(* Logix 5000 project; controller MV vendor 1 type 14 code 217 rev 31.11; software revision 31.00; part 39 of 53 *)
(* tags used below, declared in another part *)
   CWD : CHECKWORD_FLAGS;
   indirect_bit_temp : INT;
   MV_B100 : INT[255];   // AT FLAGS
   MV_MV37_AV01 : PlantItem;   // MV37_AV01
   MV_MV37_AV01_RawOutput : ALIAS FOR Remote_IO:16:O.Data.1;   // MV_MV37_AV01 MV37 coolant SOV
   MV_MV38_AV01 : PlantItem;   // MV38_AV01
   MV_MV38_AV01_RawOutput : ALIAS FOR Remote_IO:16:O.Data.2;   // MV_MV38_AV01 MV38 coolant SOV
   MV_MV39_AV01 : PlantItem;   // MV39_AV01
   MV_MV39_AV01_RawOutput : ALIAS FOR Remote_IO:16:O.Data.3;   // MV_MV39_AV01 MV39 coolant SOV
   MV_MV40_AV01 : PlantItem;   // MV40_AV01
   MV_MV40_AV01_RawOutput : ALIAS FOR Remote_IO:16:O.Data.4;   // MV_MV40_AV01 MV40 coolant SOV
   MV_MV41_AV01 : PlantItem;   // MV41_AV01
   MV_MV41_AV01_RawOutput : ALIAS FOR Remote_IO:16:O.Data.5;   // MV_MV41_AV01 MV41 coolant SOV
   MV_MV42_AV01 : PlantItem;   // MV42_AV01
   MV_MV42_AV01_RawOutput : ALIAS FOR Remote_IO:16:O.Data.6;   // MV_MV42_AV01 MV42 coolant SOV
   MV_MV43_AV01 : PlantItem;   // MV43_AV01
   MV_MV43_AV01_RawOutput : ALIAS FOR Remote_IO:16:O.Data.7;   // MV_MV43_AV01 MV43 coolant SOV
   MV_MV44_AV01 : PlantItem;   // MV44_AV01
   MV_MV44_AV01_RawOutput : ALIAS FOR Remote_IO:16:O.Data.8;   // MV_MV44_AV01 MV44 coolant SOV
   MV_MV45_AV01 : PlantItem;   // MV45_AV01
   MV_MV45_AV01_RawOutput : ALIAS FOR Remote_IO:16:O.Data.9;   // MV_MV45_AV01 MV45 coolant SOV
   MV_MV46_AV01 : PlantItem;   // MV46_AV01
   MV_MV46_AV01_RawOutput : ALIAS FOR Remote_IO:16:O.Data.10;   // MV_MV46_AV01 MV46 coolant SOV
   MV_MV47_AV01 : PlantItem;   // MV47_AV01
   MV_MV47_AV01_RawOutput : ALIAS FOR Remote_IO:16:O.Data.11;   // MV_MV47_AV01 MV47 coolant SOV
   MV_N101 : INT[255];   // AT INT Fermentation control integer workspace
   MV_N104 : INT[255];   // MV_PC_BUF PC>PLC Attemporation Control Command Buf fer File
(* MV_Common, continued *)

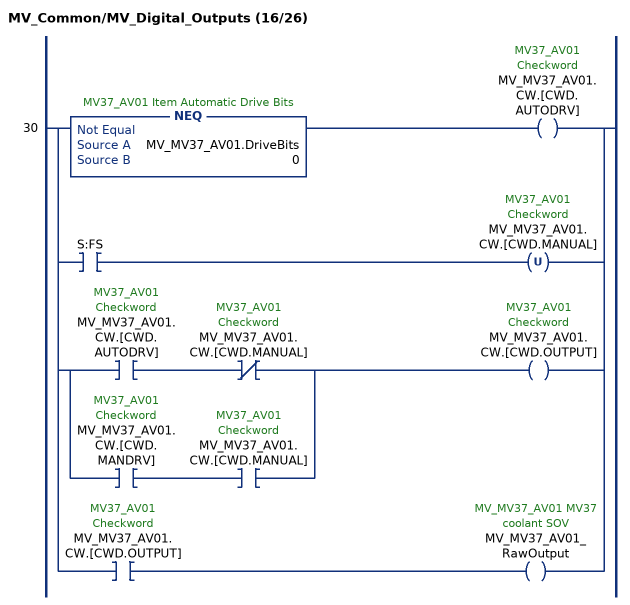
   [picture p908: MV_Common/MV_Digital_Outputs rungs 30-30]
   30: [NEQ(MV_MV37_AV01.DriveBits,0) OTE(MV_MV37_AV01.CW.[CWD.AUTODRV]) ,XIC(S:FS) OTU(MV_MV37_AV01.CW.[CWD.MANUAL]) ,[XIC(MV_MV37_AV01.CW.[CWD.AUTODRV]) XIO(MV_MV37_AV01.CW.[CWD.MANUAL]) ,XIC(MV_MV37_AV01.CW.[CWD.MANDRV]) XIC(MV_MV37_AV01.CW.[CWD.MANUAL]) ] OTE(MV_MV37_AV01.CW.[CWD.OUTPUT]) ,XIC(MV_MV37_AV01.CW.[CWD.OUTPUT]) OTE(MV_MV37_AV01_RawOutput) ];
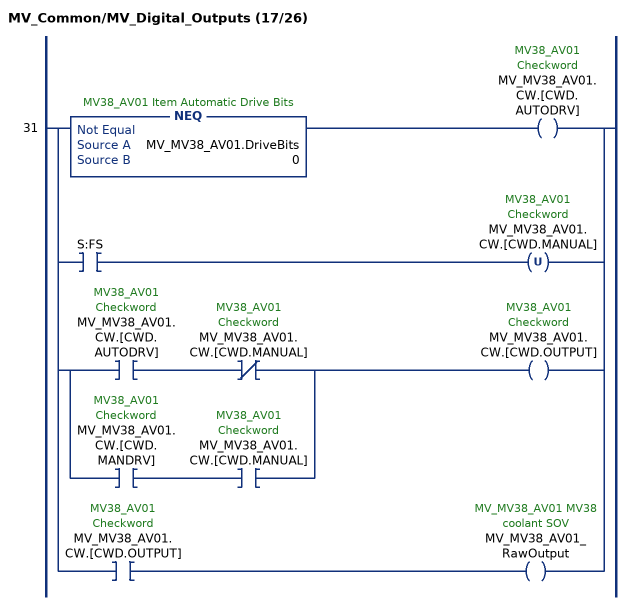
   31: [NEQ(MV_MV38_AV01.DriveBits,0) OTE(MV_MV38_AV01.CW.[CWD.AUTODRV]) ,XIC(S:FS) OTU(MV_MV38_AV01.CW.[CWD.MANUAL]) ,[XIC(MV_MV38_AV01.CW.[CWD.AUTODRV]) XIO(MV_MV38_AV01.CW.[CWD.MANUAL]) ,XIC(MV_MV38_AV01.CW.[CWD.MANDRV]) XIC(MV_MV38_AV01.CW.[CWD.MANUAL]) ] OTE(MV_MV38_AV01.CW.[CWD.OUTPUT]) ,XIC(MV_MV38_AV01.CW.[CWD.OUTPUT]) OTE(MV_MV38_AV01_RawOutput) ];
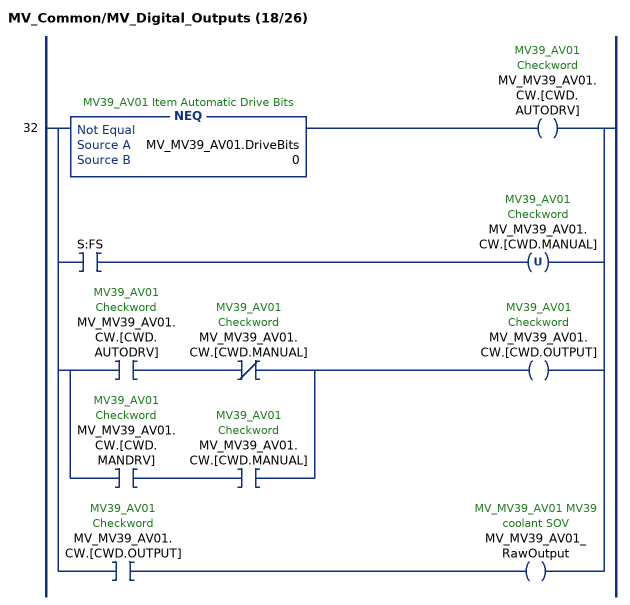
   32: [NEQ(MV_MV39_AV01.DriveBits,0) OTE(MV_MV39_AV01.CW.[CWD.AUTODRV]) ,XIC(S:FS) OTU(MV_MV39_AV01.CW.[CWD.MANUAL]) ,[XIC(MV_MV39_AV01.CW.[CWD.AUTODRV]) XIO(MV_MV39_AV01.CW.[CWD.MANUAL]) ,XIC(MV_MV39_AV01.CW.[CWD.MANDRV]) XIC(MV_MV39_AV01.CW.[CWD.MANUAL]) ] OTE(MV_MV39_AV01.CW.[CWD.OUTPUT]) ,XIC(MV_MV39_AV01.CW.[CWD.OUTPUT]) OTE(MV_MV39_AV01_RawOutput) ];
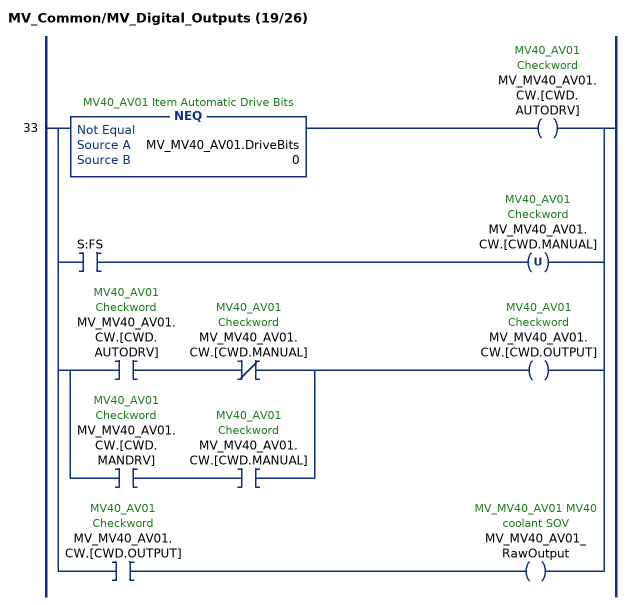
   33: [NEQ(MV_MV40_AV01.DriveBits,0) OTE(MV_MV40_AV01.CW.[CWD.AUTODRV]) ,XIC(S:FS) OTU(MV_MV40_AV01.CW.[CWD.MANUAL]) ,[XIC(MV_MV40_AV01.CW.[CWD.AUTODRV]) XIO(MV_MV40_AV01.CW.[CWD.MANUAL]) ,XIC(MV_MV40_AV01.CW.[CWD.MANDRV]) XIC(MV_MV40_AV01.CW.[CWD.MANUAL]) ] OTE(MV_MV40_AV01.CW.[CWD.OUTPUT]) ,XIC(MV_MV40_AV01.CW.[CWD.OUTPUT]) OTE(MV_MV40_AV01_RawOutput) ];
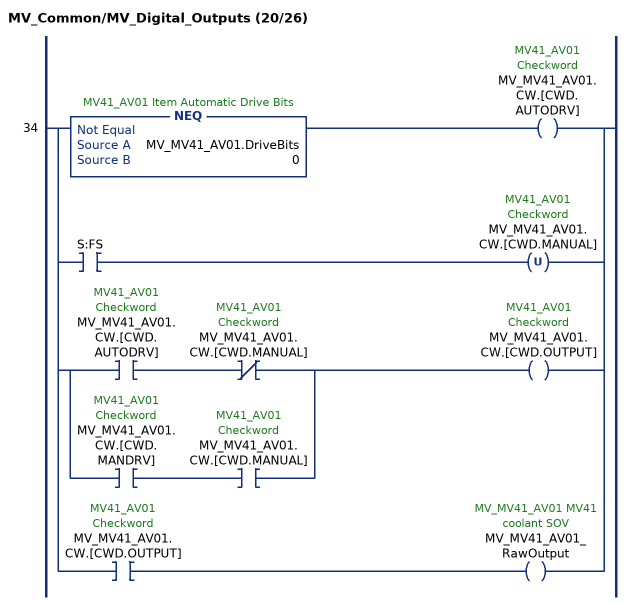
   34: [NEQ(MV_MV41_AV01.DriveBits,0) OTE(MV_MV41_AV01.CW.[CWD.AUTODRV]) ,XIC(S:FS) OTU(MV_MV41_AV01.CW.[CWD.MANUAL]) ,[XIC(MV_MV41_AV01.CW.[CWD.AUTODRV]) XIO(MV_MV41_AV01.CW.[CWD.MANUAL]) ,XIC(MV_MV41_AV01.CW.[CWD.MANDRV]) XIC(MV_MV41_AV01.CW.[CWD.MANUAL]) ] OTE(MV_MV41_AV01.CW.[CWD.OUTPUT]) ,XIC(MV_MV41_AV01.CW.[CWD.OUTPUT]) OTE(MV_MV41_AV01_RawOutput) ];
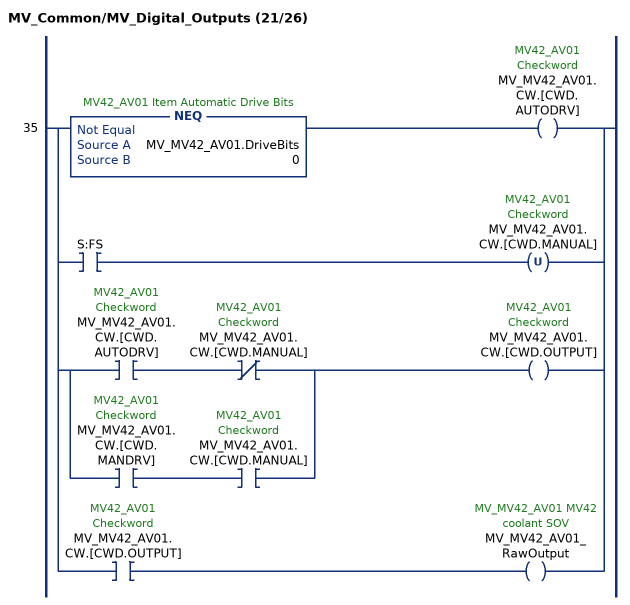
   35: [NEQ(MV_MV42_AV01.DriveBits,0) OTE(MV_MV42_AV01.CW.[CWD.AUTODRV]) ,XIC(S:FS) OTU(MV_MV42_AV01.CW.[CWD.MANUAL]) ,[XIC(MV_MV42_AV01.CW.[CWD.AUTODRV]) XIO(MV_MV42_AV01.CW.[CWD.MANUAL]) ,XIC(MV_MV42_AV01.CW.[CWD.MANDRV]) XIC(MV_MV42_AV01.CW.[CWD.MANUAL]) ] OTE(MV_MV42_AV01.CW.[CWD.OUTPUT]) ,XIC(MV_MV42_AV01.CW.[CWD.OUTPUT]) OTE(MV_MV42_AV01_RawOutput) ];
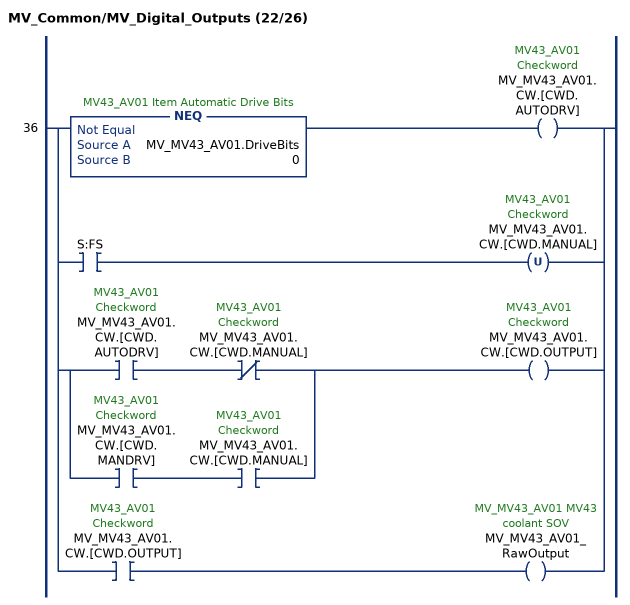
   36: [NEQ(MV_MV43_AV01.DriveBits,0) OTE(MV_MV43_AV01.CW.[CWD.AUTODRV]) ,XIC(S:FS) OTU(MV_MV43_AV01.CW.[CWD.MANUAL]) ,[XIC(MV_MV43_AV01.CW.[CWD.AUTODRV]) XIO(MV_MV43_AV01.CW.[CWD.MANUAL]) ,XIC(MV_MV43_AV01.CW.[CWD.MANDRV]) XIC(MV_MV43_AV01.CW.[CWD.MANUAL]) ] OTE(MV_MV43_AV01.CW.[CWD.OUTPUT]) ,XIC(MV_MV43_AV01.CW.[CWD.OUTPUT]) OTE(MV_MV43_AV01_RawOutput) ];
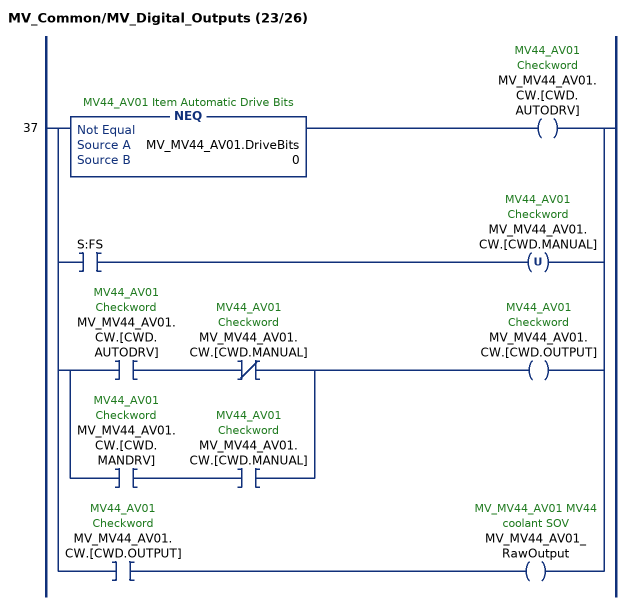
   37: [NEQ(MV_MV44_AV01.DriveBits,0) OTE(MV_MV44_AV01.CW.[CWD.AUTODRV]) ,XIC(S:FS) OTU(MV_MV44_AV01.CW.[CWD.MANUAL]) ,[XIC(MV_MV44_AV01.CW.[CWD.AUTODRV]) XIO(MV_MV44_AV01.CW.[CWD.MANUAL]) ,XIC(MV_MV44_AV01.CW.[CWD.MANDRV]) XIC(MV_MV44_AV01.CW.[CWD.MANUAL]) ] OTE(MV_MV44_AV01.CW.[CWD.OUTPUT]) ,XIC(MV_MV44_AV01.CW.[CWD.OUTPUT]) OTE(MV_MV44_AV01_RawOutput) ];
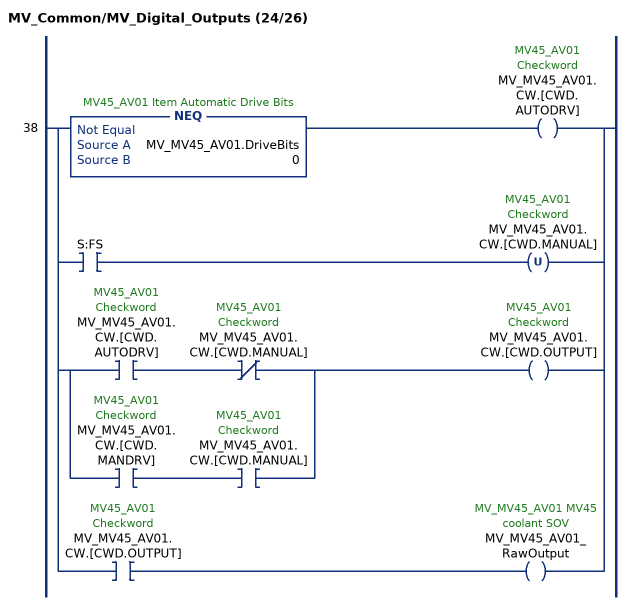
   38: [NEQ(MV_MV45_AV01.DriveBits,0) OTE(MV_MV45_AV01.CW.[CWD.AUTODRV]) ,XIC(S:FS) OTU(MV_MV45_AV01.CW.[CWD.MANUAL]) ,[XIC(MV_MV45_AV01.CW.[CWD.AUTODRV]) XIO(MV_MV45_AV01.CW.[CWD.MANUAL]) ,XIC(MV_MV45_AV01.CW.[CWD.MANDRV]) XIC(MV_MV45_AV01.CW.[CWD.MANUAL]) ] OTE(MV_MV45_AV01.CW.[CWD.OUTPUT]) ,XIC(MV_MV45_AV01.CW.[CWD.OUTPUT]) OTE(MV_MV45_AV01_RawOutput) ];
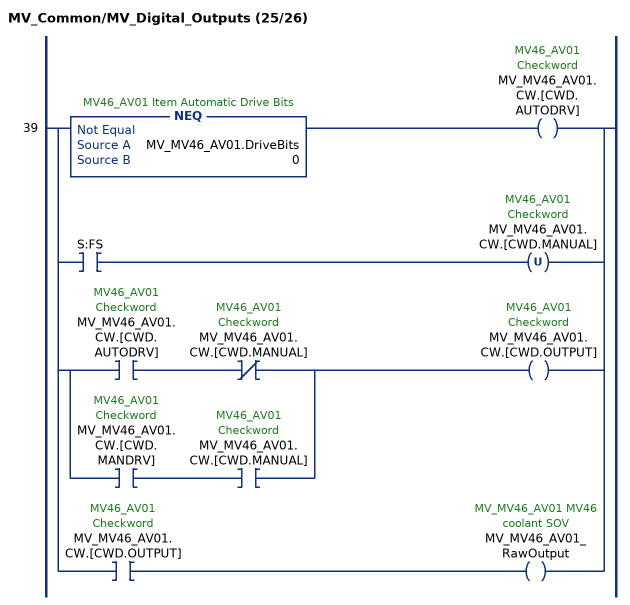
   39: [NEQ(MV_MV46_AV01.DriveBits,0) OTE(MV_MV46_AV01.CW.[CWD.AUTODRV]) ,XIC(S:FS) OTU(MV_MV46_AV01.CW.[CWD.MANUAL]) ,[XIC(MV_MV46_AV01.CW.[CWD.AUTODRV]) XIO(MV_MV46_AV01.CW.[CWD.MANUAL]) ,XIC(MV_MV46_AV01.CW.[CWD.MANDRV]) XIC(MV_MV46_AV01.CW.[CWD.MANUAL]) ] OTE(MV_MV46_AV01.CW.[CWD.OUTPUT]) ,XIC(MV_MV46_AV01.CW.[CWD.OUTPUT]) OTE(MV_MV46_AV01_RawOutput) ];
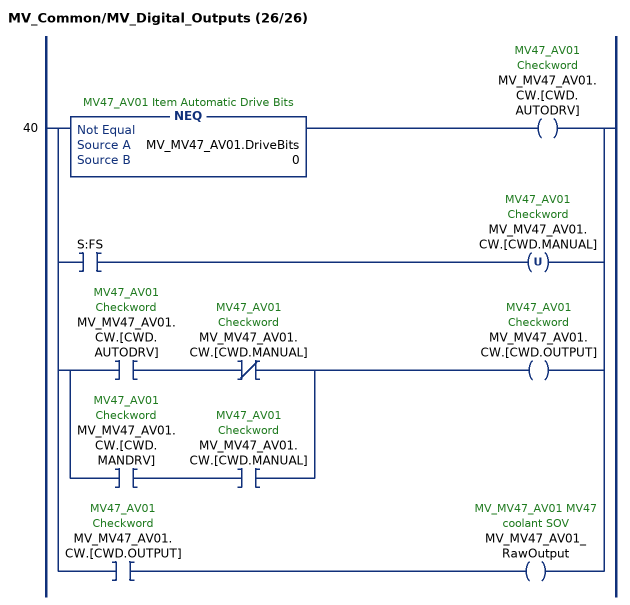
   40: [NEQ(MV_MV47_AV01.DriveBits,0) OTE(MV_MV47_AV01.CW.[CWD.AUTODRV]) ,XIC(S:FS) OTU(MV_MV47_AV01.CW.[CWD.MANUAL]) ,[XIC(MV_MV47_AV01.CW.[CWD.AUTODRV]) XIO(MV_MV47_AV01.CW.[CWD.MANUAL]) ,XIC(MV_MV47_AV01.CW.[CWD.MANDRV]) XIC(MV_MV47_AV01.CW.[CWD.MANUAL]) ] OTE(MV_MV47_AV01.CW.[CWD.OUTPUT]) ,XIC(MV_MV47_AV01.CW.[CWD.OUTPUT]) OTE(MV_MV47_AV01_RawOutput) ];
END_ROUTINE

ROUTINE MV_FV_COMMAND_101   (* ladder *)
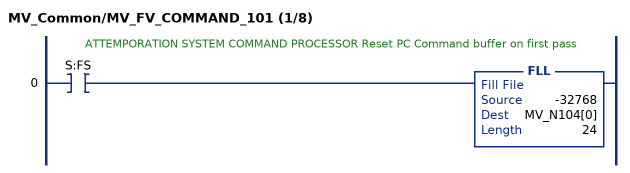
   // ATTEMPORATION SYSTEM COMMAND PROCESSOR Reset PC Command buffer on first pass
   0: XIC(S:FS)FLL(-32768,MV_N104[0],24);
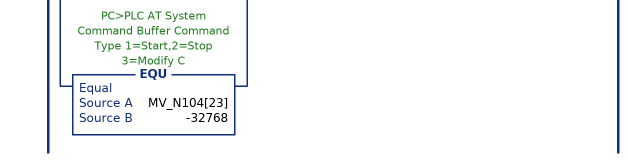
   // WAIT FOR PC TO SEND NEW COMMAND If any word within the PC/PLC system command buffer contains -32768, the block has not yet been fully downloaded and therefore no new command has been requested.
   1: [EQU(MV_N104[0],-32768) ,EQU(MV_N104[1],-32768) ,EQU(MV_N104[2],-32768) ,EQU(MV_N104[3],-32768) ,EQU(MV_N104[4],-32768) ,EQU(MV_N104[5],-32768) ,EQU(MV_N104[6],-32768) ,EQU(MV_N104[7],-32768) ,EQU(MV_N104[8],-32768) ,EQU(MV_N104[9],-32768) ,EQU(MV_N104[10],-32768) ,EQU(MV_N104[11],-32768) ,EQU(MV_N104[12],-32768) ,EQU(MV_N104[13],-32768) ,EQU(MV_N104[14],-32768) ,EQU(MV_N104[15],-32768) ,EQU(MV_N104[16],-32768) ,EQU(MV_N104[17],-32768) ,EQU(MV_N104[18],-32768) ,EQU(MV_N104[19],-32768) ,EQU(MV_N104[20],-32768) ,EQU(MV_N104[21],-32768) ,EQU(MV_N104[22],-32768) ,EQU(MV_N104[23],-32768) ]OTE(MV_B100[1].0);
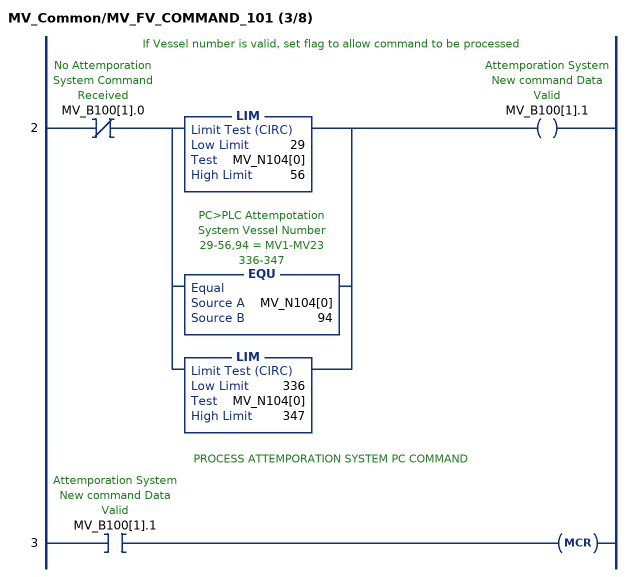
   // If Vessel number is valid, set flag to allow command to be processed
   2: XIO(MV_B100[1].0)[LIM(29,MV_N104[0],56) ,EQU(MV_N104[0],94) ,LIM(336,MV_N104[0],347) ]OTE(MV_B100[1].1);
   // PROCESS ATTEMPORATION SYSTEM PC COMMAND
   3: XIC(MV_B100[1].1)MCR();
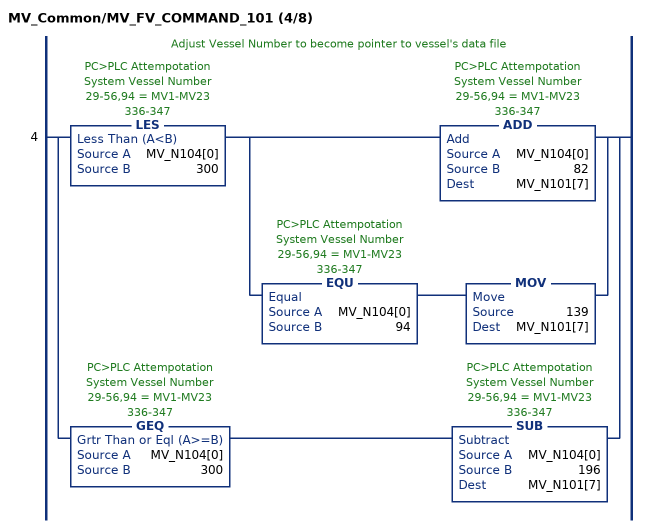
   // Adjust Vessel Number to become pointer to vessel's data file
   4: [LES(MV_N104[0],300) [ADD(MV_N104[0],82,MV_N101[7]) ,EQU(MV_N104[0],94) MOV(139,MV_N101[7]) ] ,GEQ(MV_N104[0],300) SUB(MV_N104[0],196,MV_N101[7]) ];
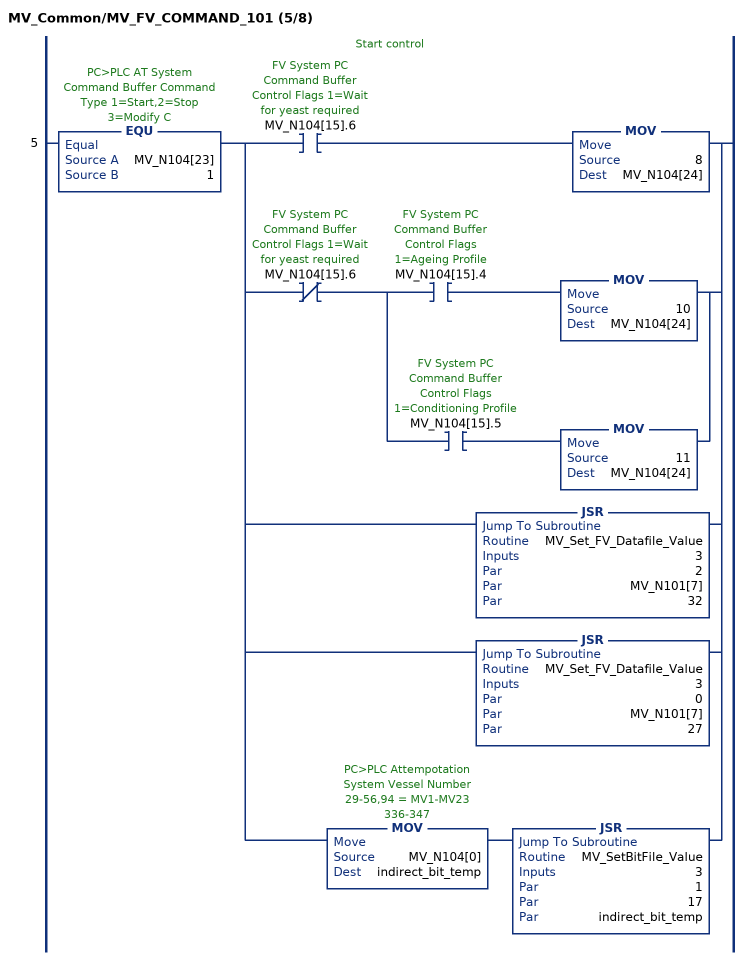
   // Start control
   5: EQU(MV_N104[23],1)[XIC(MV_N104[15].6) MOV(8,MV_N104[24]) ,XIO(MV_N104[15].6) [XIC(MV_N104[15].4) MOV(10,MV_N104[24]) ,XIC(MV_N104[15].5) MOV(11,MV_N104[24]) ] ,JSR(MV_Set_FV_Datafile_Value,3,2,MV_N101[7],32) ,JSR(MV_Set_FV_Datafile_Value,3,0,MV_N101[7],27) ,MOV(MV_N104[0],indirect_bit_temp) JSR(MV_SetBitFile_Value,3,1,17,indirect_bit_temp) ];
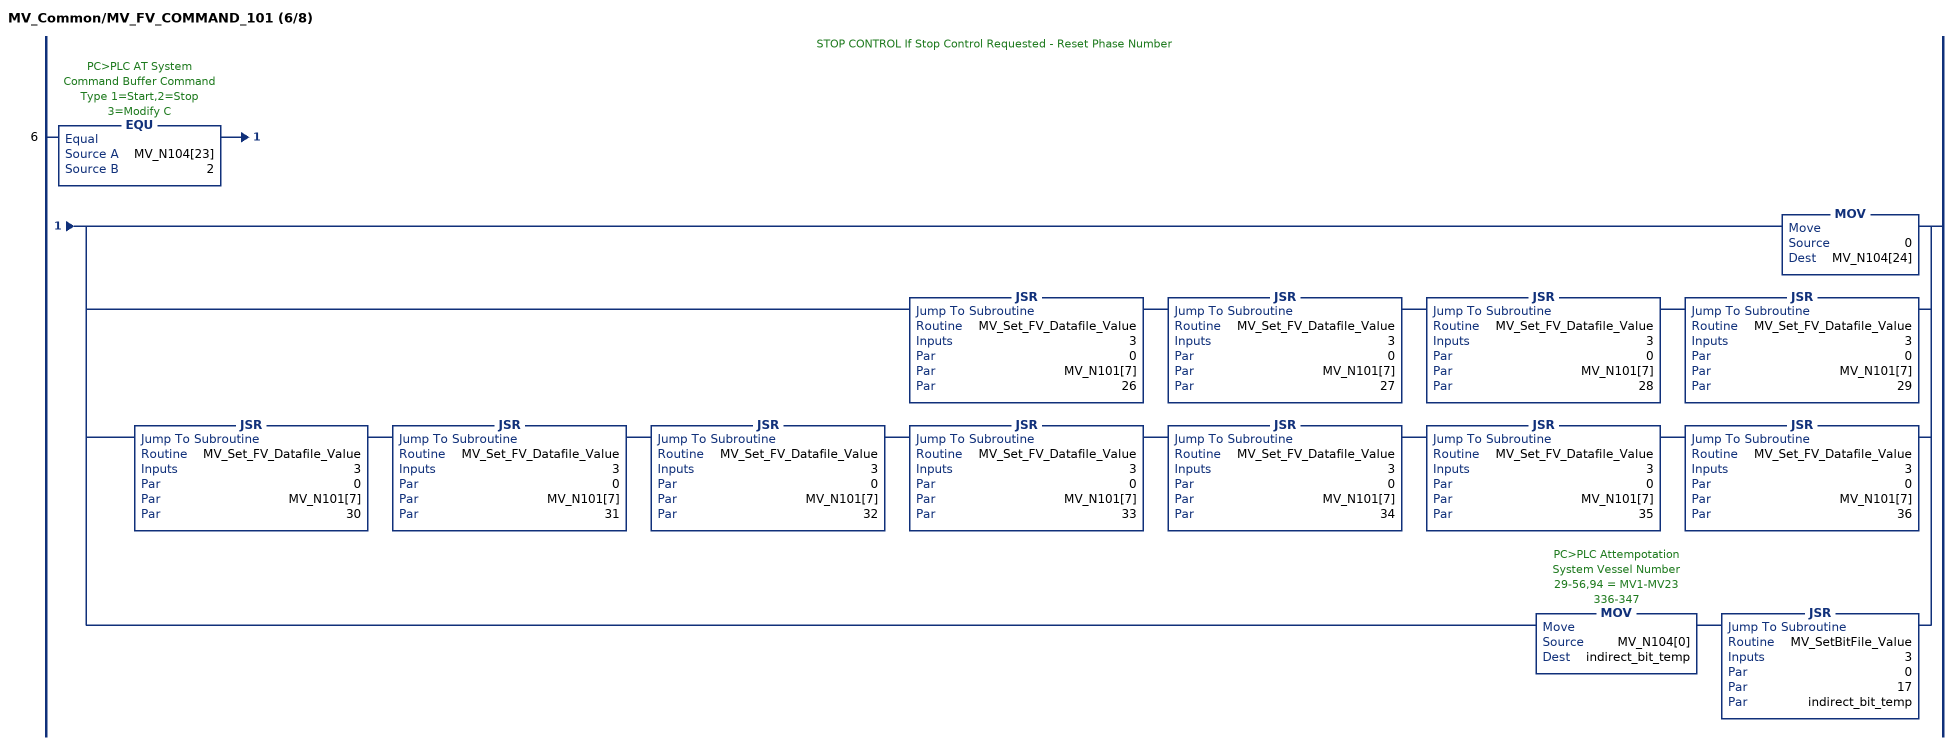
   // STOP CONTROL If Stop Control Requested - Reset Phase Number
   6: EQU(MV_N104[23],2)[MOV(0,MV_N104[24]) ,JSR(MV_Set_FV_Datafile_Value,3,0,MV_N101[7],26) JSR(MV_Set_FV_Datafile_Value,3,0,MV_N101[7],27) JSR(MV_Set_FV_Datafile_Value,3,0,MV_N101[7],28) JSR(MV_Set_FV_Datafile_Value,3,0,MV_N101[7],29) ,JSR(MV_Set_FV_Datafile_Value,3,0,MV_N101[7],30) JSR(MV_Set_FV_Datafile_Value,3,0,MV_N101[7],31) JSR(MV_Set_FV_Datafile_Value,3,0,MV_N101[7],32) JSR(MV_Set_FV_Datafile_Value,3,0,MV_N101[7],33) JSR(MV_Set_FV_Datafile_Value,3,0,MV_N101[7],34) JSR(MV_Set_FV_Datafile_Value,3,0,MV_N101[7],35) JSR(MV_Set_FV_Datafile_Value,3,0,MV_N101[7],36) ,MOV(MV_N104[0],indirect_bit_temp) JSR(MV_SetBitFile_Value,3,0,17,indirect_bit_temp) ];
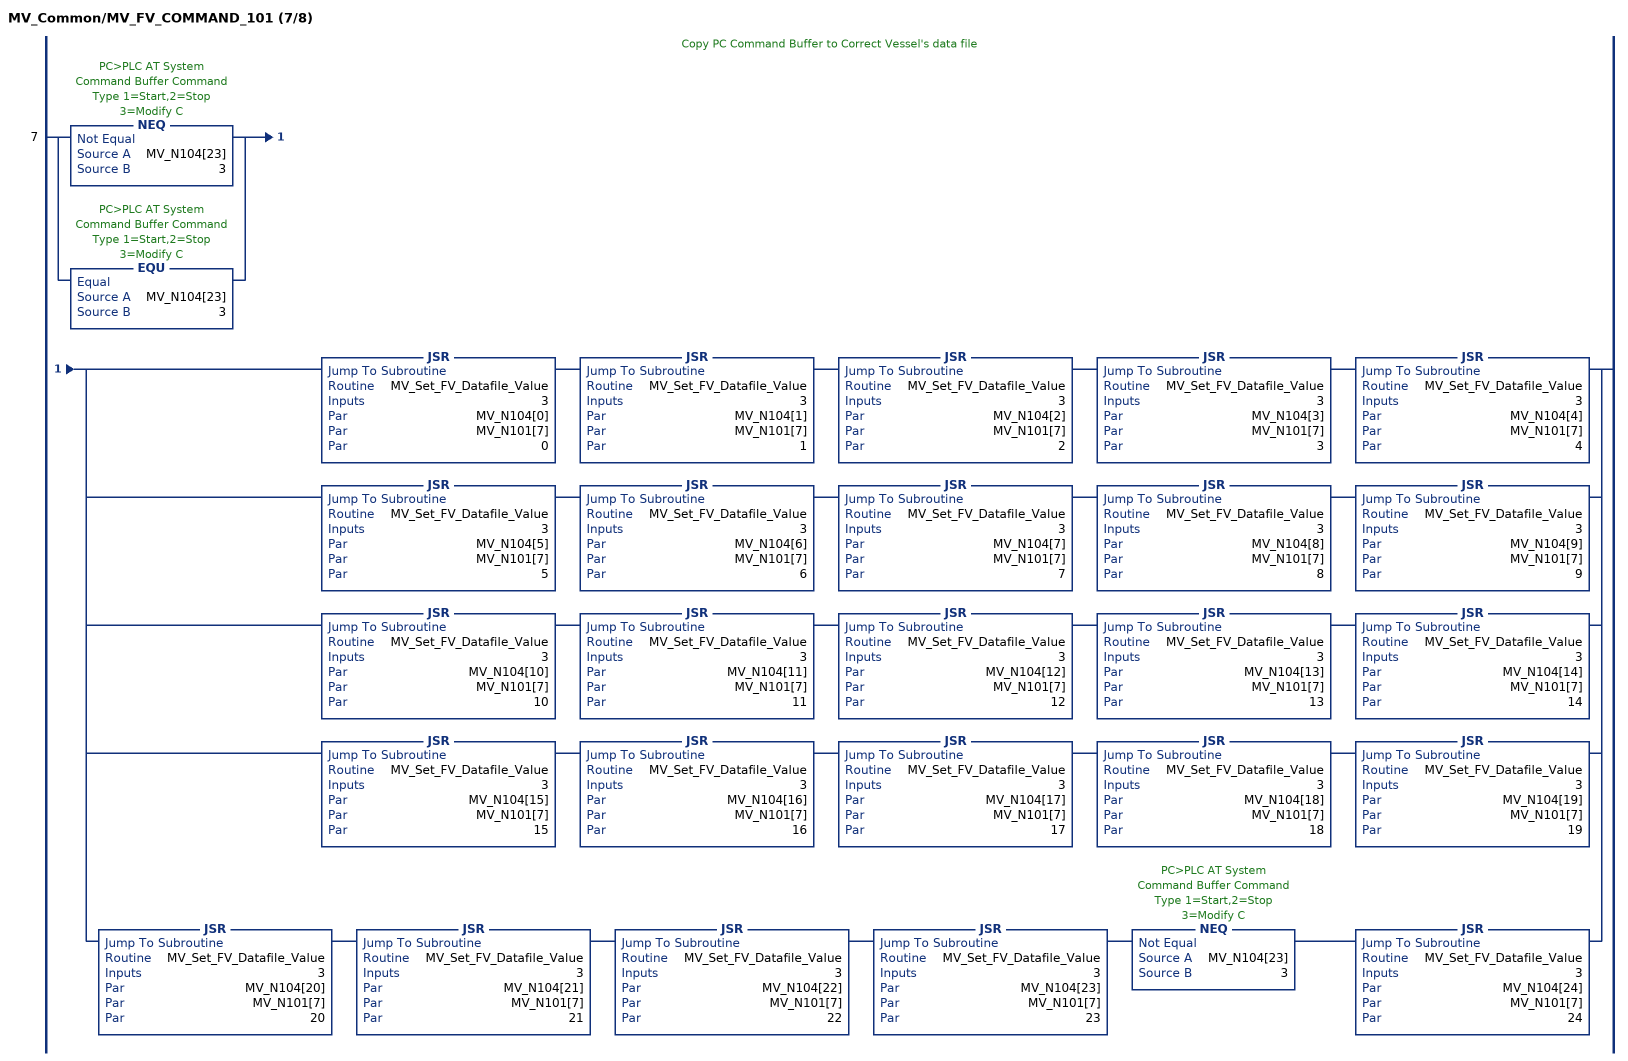
   // Copy PC Command Buffer to Correct Vessel's data file
   7: [NEQ(MV_N104[23],3) ,EQU(MV_N104[23],3) ][JSR(MV_Set_FV_Datafile_Value,3,MV_N104[0],MV_N101[7],0) JSR(MV_Set_FV_Datafile_Value,3,MV_N104[1],MV_N101[7],1) JSR(MV_Set_FV_Datafile_Value,3,MV_N104[2],MV_N101[7],2) JSR(MV_Set_FV_Datafile_Value,3,MV_N104[3],MV_N101[7],3) JSR(MV_Set_FV_Datafile_Value,3,MV_N104[4],MV_N101[7],4) ,JSR(MV_Set_FV_Datafile_Value,3,MV_N104[5],MV_N101[7],5) JSR(MV_Set_FV_Datafile_Value,3,MV_N104[6],MV_N101[7],6) JSR(MV_Set_FV_Datafile_Value,3,MV_N104[7],MV_N101[7],7) JSR(MV_Set_FV_Datafile_Value,3,MV_N104[8],MV_N101[7],8) JSR(MV_Set_FV_Datafile_Value,3,MV_N104[9],MV_N101[7],9) ,JSR(MV_Set_FV_Datafile_Value,3,MV_N104[10],MV_N101[7],10) JSR(MV_Set_FV_Datafile_Value,3,MV_N104[11],MV_N101[7],11) JSR(MV_Set_FV_Datafile_Value,3,MV_N104[12],MV_N101[7],12) JSR(MV_Set_FV_Datafile_Value,3,MV_N104[13],MV_N101[7],13) JSR(MV_Set_FV_Datafile_Value,3,MV_N104[14],MV_N101[7],14) ,JSR(MV_Set_FV_Datafile_Value,3,MV_N104[15],MV_N101[7],15) JSR(MV_Set_FV_Datafile_Value,3,MV_N104[16],MV_N101[7],16) JSR(MV_Set_FV_Datafile_Value,3,MV_N104[17],MV_N101[7],17) JSR(MV_Set_FV_Datafile_Value,3,MV_N104[18],MV_N101[7],18) JSR(MV_Set_FV_Datafile_Value,3,MV_N104[19],MV_N101[7],19) ,JSR(MV_Set_FV_Datafile_Value,3,MV_N104[20],MV_N101[7],20) JSR(MV_Set_FV_Datafile_Value,3,MV_N104[21],MV_N101[7],21) JSR(MV_Set_FV_Datafile_Value,3,MV_N104[22],MV_N101[7],22) JSR(MV_Set_FV_Datafile_Value,3,MV_N104[23],MV_N101[7],23) NEQ(MV_N104[23],3) JSR(MV_Set_FV_Datafile_Value,3,MV_N104[24],MV_N101[7],24) ];
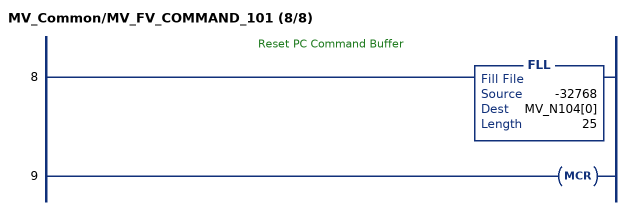
   // Reset PC Command Buffer
   8: FLL(-32768,MV_N104[0],25);
   9: MCR();
END_ROUTINE
